HMI tags "Standard-Variablentabelle"
   "Trigger" : Int, internal
   "TP_Online" : Int, internal
   "_BildNr_aktuell" : Int, internal
   "__Pult_Name" : Int, internal
   "__Pult_Name(1)" : WString[10], internal
   "test" : Int, internal
   "LinePLC1_RD_ready" : Bool = PLC LinePLC1_RD_ready AT %I4248.0, 1 s
   "DiagStatusUpdate" : Bool = PLC DiagStatusUpdate AT %M1.1, 1 s
   "EMS_Carrier_Spacing" : Int = PLC EMS.Carrier_Spacing, 1 s
   "EMS_Coarse_Decel_Speed" : Word = PLC EMS.CoarseDecelSpeed AT %DB1.DBW0, 1 s
   "EMS_Coarse_Position_Decel_Offset" : Word = PLC EMS.CoarsePositionDecelOffset AT %DB1.DBW0, 1 s
   "EMS_Coarse_Position_Tolerance" : Word = PLC EMS.CoarsePositionTolerance AT %DB1.DBW0, 1 s
   "EMS_Fine_Decel_Speed" : Word = PLC EMS.FineDecelSpeed AT %DB1.DBW0, 1 s
   "EMS_Fine_Posistion_Tolerance" : Word = PLC EMS.FinePositionTolerance AT %DB1.DBW0, 1 s
   "EMS_Fine_Position_Decel_Offset" : Word = PLC EMS.FinePositionDecelOffset AT %DB1.DBW0, 1 s
   "EMS_Production_Spacing" : Word = PLC EMS.Production_Spacing, 1 s
   "EMS_Production_Zone_Speed" : Word = PLC EMS.ProductionZnSpeed AT %DB1.DBW0, 1 s
   "Temp_Placeholder" : Int = PLC Temp_Int AT %MW56, 1 s
   "CARRIER #01   CURRENT" : Int = PLC "CARRIER #01   CURRENT" AT %MW72, 1 s
   "CARRIER #01   G120D Status WORD.0(1)" : Bool = PLC "CARRIER #01   G120D STATUS WORD.0" AT %M76.0, 1 s
   "CARRIER #01   G120D Status WORD.1(1)" : Bool = PLC "CARRIER #01   G120D STATUS WORD.1" AT %M76.1, 1 s
   "CARRIER #01   G120D Status WORD.10(1)" : Bool = PLC "CARRIER #01   G120D STATUS WORD.10" AT %M77.2, 1 s
   "CARRIER #01   G120D Status WORD.11(1)" : Bool = PLC "CARRIER #01   G120D STATUS WORD.11" AT %M77.3, 1 s
   "CARRIER #01   G120D Status WORD.12(1)" : Bool = PLC "CARRIER #01   G120D STATUS WORD.12" AT %M77.4, 1 s
   "CARRIER #01   G120D Status WORD.13(1)" : Bool = PLC "CARRIER #01   G120D STATUS WORD.13" AT %M77.5, 1 s
   "CARRIER #01   G120D Status WORD.14(1)" : Bool = PLC "CARRIER #01   G120D STATUS WORD.14" AT %M77.6, 1 s
   "CARRIER #01   G120D Status WORD.15(1)" : Bool = PLC "CARRIER #01   G120D STATUS WORD.15" AT %M77.7, 1 s
   "CARRIER #01   G120D Status WORD.2(1)" : Bool = PLC "CARRIER #01   G120D STATUS WORD.2" AT %M76.2, 1 s
   "CARRIER #01   G120D Status WORD.3(1)" : Bool = PLC "CARRIER #01   G120D STATUS WORD.3" AT %M76.3, 1 s
   "CARRIER #01   G120D Status WORD.4(1)" : Bool = PLC "CARRIER #01   G120D STATUS WORD.4" AT %M76.4, 1 s
   "CARRIER #01   G120D Status WORD.5(1)" : Bool = PLC "CARRIER #01   G120D STATUS WORD.5" AT %M76.5, 1 s
   "CARRIER #01   G120D Status WORD.6(1)" : Bool = PLC "CARRIER #01   G120D STATUS WORD.6" AT %M76.6, 1 s
   "CARRIER #01   G120D Status WORD.7(1)" : Bool = PLC "CARRIER #01   G120D STATUS WORD.7" AT %M76.7, 1 s
   "CARRIER #01   G120D Status WORD.8(1)" : Bool = PLC "CARRIER #01   G120D STATUS WORD.8" AT %M77.0, 1 s
   "CARRIER #01   G120D Status WORD.9(1)" : Bool = PLC "CARRIER #01   G120D STATUS WORD.9" AT %M77.1, 1 s
   "CARRIER #01   G120D STATUS WORD.0" : Bool = PLC "CARRIER #01   G120D STATUS WORD.0" AT %M76.0, 1 s
   "CARRIER #01   G120D STATUS WORD.1" : Bool = PLC "CARRIER #01   G120D STATUS WORD.1" AT %M76.1, 1 s
   "CARRIER #01   G120D STATUS WORD.10" : Bool = PLC "CARRIER #01   G120D STATUS WORD.10" AT %M77.2, 1 s
   "CARRIER #01   G120D STATUS WORD.11" : Bool = PLC "CARRIER #01   G120D STATUS WORD.11" AT %M77.3, 1 s
   "CARRIER #01   G120D STATUS WORD.12" : Bool = PLC "CARRIER #01   G120D STATUS WORD.12" AT %M77.4, 1 s
   "CARRIER #01   G120D STATUS WORD.13" : Bool = PLC "CARRIER #01   G120D STATUS WORD.13" AT %M77.5, 1 s
   "CARRIER #01   G120D STATUS WORD.14" : Bool = PLC "CARRIER #01   G120D STATUS WORD.14" AT %M77.6, 1 s
   "CARRIER #01   G120D STATUS WORD.15" : Bool = PLC "CARRIER #01   G120D STATUS WORD.15" AT %M77.7, 1 s
   "CARRIER #01   G120D STATUS WORD.2" : Bool = PLC "CARRIER #01   G120D STATUS WORD.2" AT %M76.2, 1 s
   "CARRIER #01   G120D STATUS WORD.3" : Bool = PLC "CARRIER #01   G120D STATUS WORD.3" AT %M76.3, 1 s
   "CARRIER #01   G120D STATUS WORD.4" : Bool = PLC "CARRIER #01   G120D STATUS WORD.4" AT %M76.4, 1 s
   "CARRIER #01   G120D STATUS WORD.5" : Bool = PLC "CARRIER #01   G120D STATUS WORD.5" AT %M76.5, 1 s
   "CARRIER #01   G120D STATUS WORD.6" : Bool = PLC "CARRIER #01   G120D STATUS WORD.6" AT %M76.6, 1 s
   "CARRIER #01   G120D STATUS WORD.7" : Bool = PLC "CARRIER #01   G120D STATUS WORD.7" AT %M76.7, 1 s
   "CARRIER #01   G120D STATUS WORD.8" : Bool = PLC "CARRIER #01   G120D STATUS WORD.8" AT %M77.0, 1 s
   "CARRIER #01   G120D STATUS WORD.9" : Bool = PLC "CARRIER #01   G120D STATUS WORD.9" AT %M77.1, 1 s
   "CARRIER #01   POSITION" : Int = PLC "CARRIER #01   POSITION" AT %MW78, 1 s
   "CARRIER #01 480VPowerOn_MDCB1" : Bool = PLC "CARRIER #01 480VPowerOn_MDCB1" AT %M80.0, 1 s
   "CARRIER #01 CrashDetectSW" : Bool = PLC "CARRIER #01 CrashDetectSW" AT %M80.1, 1 s
   "CARRIER #01 DCsupplyOnPSCB2" : Bool = PLC "CARRIER #01 DCsupplyOnPSCB2" AT %M80.2, 1 s
   "CARRIER #01 FaultLight_LH" : Bool = PLC "CARRIER #01 FaultLight_LH" AT %M80.3, 1 s
   "CARRIER #01 FaultLight_RH" : Bool = PLC "CARRIER #01 FaultLight_RH" AT %M80.4, 1 s
   "Carrier #01 HMI 1 Status0.5(1)" : Bool = PLC "CARRIER #01   1 STATUS [0].5" AT %M80.5, 1 s
   "CARRIER #01 PB1_ProdHoldLH" : Bool = PLC "CARRIER #01 PB1_ProdHoldLH" AT %M80.6, 1 s
   "CARRIER #01 PB2_ResetLH" : Bool = PLC "CARRIER #01 PB2_ResetLH" AT %M80.7, 1 s
   "CARRIER #01 PB3_ProdHoldRH" : Bool = PLC "CARRIER #01 PB3_ProdHoldRH" AT %M81.0, 1 s
   "CARRIER #01 PB4_ResetRH" : Bool = PLC "CARRIER #01 PB4_ResetRH" AT %M81.1, 1 s
   "CARRIER #01 RunLight_LH" : Bool = PLC "CARRIER #01 RunLight_LH" AT %M81.2, 1 s
   "CARRIER #01 RunLight_RH" : Bool = PLC "CARRIER #01 RunLight_RH" AT %M81.3, 1 s
   "CARRIER #01 SitopSelectStatus" : Bool = PLC "CARRIER #01 SitopSelectStatus" AT %M81.4, 1 s
   "CARRIER #01 SpareInput(2_1)" : Bool = PLC "CARRIER #01 SpareInput(2_1)" AT %M81.5, 1 s
   "CARRIER #01 SpareInput(2_2)" : Bool = PLC "CARRIER #01 SpareInput(2_2)" AT %M81.6, 1 s
   "CARRIER #01 SpareInput(2_3)" : Bool = PLC "CARRIER #01 SpareInput(2_3)" AT %M81.7, 1 s
   "CARRIER #01 SpareInput(2_4)" : Bool = PLC "CARRIER #01 SpareInput(2_4)" AT %M82.0, 1 s
   "CARRIER #01 SpareInput(2_5)" : Bool = PLC "CARRIER #01 SpareInput(2_5)" AT %M82.1, 1 s
   "CARRIER #01 SpareInput(2_6)" : Bool = PLC "CARRIER #01 SpareInput(2_6)" AT %M82.2, 1 s
   "CARRIER #01 SpareInput(2_7)" : Bool = PLC "CARRIER #01 SpareInput(2_7)" AT %M82.3, 1 s
   "CARRIER #01 SpareInput(4_1)" : Bool = PLC "CARRIER #01 SpareInput(4_1)" AT %M82.4, 1 s
   "CARRIER #01 SpareInput(4_14)" : Bool = PLC "CARRIER #01 SpareInput(4_14)" AT %M82.5, 1 s
   "CARRIER #01 SpareInput(4_15)" : Bool = PLC "CARRIER #01 SpareInput(4_15)" AT %M82.6, 1 s
   "CARRIER #01 SpareInput(4_16)" : Bool = PLC "CARRIER #01 SpareInput(4_16)" AT %M82.7, 1 s
   "CARRIER #01 SpareInput(4_17)" : Bool = PLC "CARRIER #01 SpareInput(4_17)" AT %M83.0, 1 s
   "CARRIER #01 SpareInput(4_2)" : Bool = PLC "CARRIER #01 SpareInput(4_2)" AT %M83.1, 1 s
   "CARRIER #01 SpareInput(4_5)" : Bool = PLC "CARRIER #01 SpareInput(4_5)" AT %M83.2, 1 s
   "CARRIER #01 SpareInput(4_6)" : Bool = PLC "CARRIER #01 SpareInput(4_6)" AT %M83.3, 1 s
   "CARRIER #01 SpareInput(4_7)" : Bool = PLC "CARRIER #01 SpareInput(4_7)" AT %M83.4, 1 s
   "CARRIER #01 SpareOutput(5_5)" : Bool = PLC "CARRIER #01 SpareOutput(5_5)" AT %M83.5, 1 s
   "CARRIER #01 SpareOutput(5_6)" : Bool = PLC "CARRIER #01 SpareOutput(5_6)" AT %M83.6, 1 s
   "CARRIER #01 SpareOutput(5_7)" : Bool = PLC "CARRIER #01 SpareOutput(5_7)" AT %M83.7, 1 s
   "CARRIER #01 SpareSafetyOutput(3_1)" : Bool = PLC "CARRIER #01 SpareSafetyOutput(3_1)" AT %M84.0, 1 s
   "CARRIER #01 SpareSafetyOutput(3_2)" : Bool = PLC "CARRIER #01 SpareSafetyOutput(3_2)" AT %M84.1, 1 s
   "CARRIER #01 SpareSafetyOutput(3_3)" : Bool = PLC "CARRIER #01 SpareSafetyOutput(3_3)" AT %M84.2, 1 s
   "CARRIER #01 SpareSafetyOutput(3_4)" : Bool = PLC "CARRIER #01 SpareSafetyOutput(3_4)" AT %M84.3, 1 s
   "CARRIER #01 SpareSafetyOutput(3_5)" : Bool = PLC "CARRIER #01 SpareSafetyOutput(3_5)" AT %M84.4, 1 s
   "CARRIER #01 SpareSafetyOutput(3_6)" : Bool = PLC "CARRIER #01 SpareSafetyOutput(3_6)" AT %M84.5, 1 s
   "CARRIER #01 SpareSafetyOutput(3_7)" : Bool = PLC "CARRIER #01 SpareSafetyOutput(3_7)" AT %M84.6, 1 s
   "Carrier #01_ At Command Position" : Bool = PLC DB_SDC_ERRORS_STAT.ER_AKT[49].ER_STAT[1].ERROR AT %M84.7, 1 s
   "Carrier #01_ Carrier in zone" : Int = PLC "Carrier #01_ Carrier in zone" AT %MW86, 1 s
   "Carrier #01_ Next carrier number" : Int = PLC "Carrier #01_ Next carrier number" AT %MW88, 1 s
   "Carrier 1 G120 D Status" : Bool = PLC EMS.Carrier[12].SDC_IN.DriveCommFault AT %I412.1, 1 s
   "Carrier 1 HMI Status" : Bool = PLC "Carrier 1 HMI Status" AT %I412.2, 1 s
   "Carrier 1 PnF Encoder Status" : Bool = PLC "Carrier 1 PnF Encoder Status" AT %I412.0, 1 s
   "Carrier 2  HMI Staus" : Bool = PLC "Carrier 2 HMI Status" AT %I432.2, 1 s
   "Carrier 2 G120 D Status" : Bool = PLC "Carrier 2  Drive Status" AT %I432.1, 1 s
   "Carrier 2 PnF Encoder Status" : Bool = PLC "Carrier 2 PnF Encoder Status" AT %I432.0, 1 s
   "Carrier 3  G120 D Status" : Bool = PLC "Carrier 3  Drive Status" AT %I452.1, 1 s
   "Carrier 3  PnF Encoder Status" : Bool = PLC "Carrier 3 PnF Encoder Status" AT %I452.0, 1 s
   "Carrier 3 HMI Status" : Bool = PLC "Carrier 3 HMI Status" AT %I452.2, 1 s
   "Carrier 4 G120 D Status" : Bool = PLC "Carrier 4  Drive Status" AT %I472.1, 1 s
   "Carrier 4 HMI Status" : Bool = PLC "Carrier 4 HMI Status" AT %I472.2, 1 s
   "Carrier 4 PnF Encoder Status" : Bool = PLC "Carrier 4 PnF Encoder Status" AT %I472.0, 1 s
   "Carrier_Index_HMI" : Int = PLC Carrier_Index_HMI AT %MW70, 1 s
   "Always_OFF_HMI" : Bool, internal
   "Always_ON_HMI" : Bool, internal
   "EMS_Accum_Zone_Speed" : Word = PLC EMS.AccumZnSpeed AT %DB1.DBW0, 1 s
   "PLC_IP_Address" : WString[30], internal
   "DB302_HMI_Faults_Carrier1_Faults_0" : Int = PLC DB302_HMI_Faults.Carrier1_Faults_0 AT %DB1.DBW0, 1 s
   "DB302_HMI_Faults_Carrier1_Faults_1" : Int = PLC DB302_HMI_Faults.Carrier1_Faults_1 AT %DB1.DBW0, 1 s
   "DB302_HMI_Faults_Carrier1_Faults_2" : Int = PLC DB302_HMI_Faults.Carrier1_Faults_2 AT %DB1.DBW0, 1 s
   "DB302_HMI_Faults_Carrier1_Faults_3" : Int = PLC DB302_HMI_Faults.Carrier1_Faults_3 AT %DB1.DBW0, 1 s
   "DB302_HMI_Faults_Carrier10_Faults_0" : Int = PLC DB302_HMI_Faults.Carrier10_Faults_0 AT %DB1.DBW0, 1 s
   "DB302_HMI_Faults_Carrier10_Faults_1" : Int = PLC DB302_HMI_Faults.Carrier10_Faults_1 AT %DB1.DBW0, 1 s
   "DB302_HMI_Faults_Carrier10_Faults_2" : Int = PLC DB302_HMI_Faults.Carrier10_Faults_2 AT %DB1.DBW0, 1 s
   "DB302_HMI_Faults_Carrier10_Faults_3" : Int = PLC DB302_HMI_Faults.Carrier10_Faults_3 AT %DB1.DBW0, 1 s
   "DB302_HMI_Faults_Carrier11_Faults_0" : Int = PLC DB302_HMI_Faults.Carrier11_Faults_0 AT %DB1.DBW0, 1 s
   "DB302_HMI_Faults_Carrier11_Faults_1" : Int = PLC DB302_HMI_Faults.Carrier11_Faults_1 AT %DB1.DBW0, 1 s
   "DB302_HMI_Faults_Carrier11_Faults_2" : Int = PLC DB302_HMI_Faults.Carrier11_Faults_2 AT %DB1.DBW0, 1 s
   "DB302_HMI_Faults_Carrier11_Faults_3" : Int = PLC DB302_HMI_Faults.Carrier11_Faults_3 AT %DB1.DBW0, 1 s
   "DB302_HMI_Faults_Carrier12_Faults_0" : Int = PLC DB302_HMI_Faults.Carrier12_Faults_0 AT %DB1.DBW0, 1 s
   "DB302_HMI_Faults_Carrier12_Faults_1" : Int = PLC DB302_HMI_Faults.Carrier12_Faults_1 AT %DB1.DBW0, 1 s
   "DB302_HMI_Faults_Carrier12_Faults_2" : Int = PLC DB302_HMI_Faults.Carrier12_Faults_2 AT %DB1.DBW0, 1 s
   "DB302_HMI_Faults_Carrier12_Faults_3" : Int = PLC DB302_HMI_Faults.Carrier12_Faults_3 AT %DB1.DBW0, 1 s
   "DB302_HMI_Faults_Carrier13_Faults_0" : Int = PLC DB302_HMI_Faults.Carrier13_Faults_0 AT %DB1.DBW0, 1 s
   "DB302_HMI_Faults_Carrier13_Faults_1" : Int = PLC DB302_HMI_Faults.Carrier13_Faults_1 AT %DB1.DBW0, 1 s
   "DB302_HMI_Faults_Carrier13_Faults_2" : Int = PLC DB302_HMI_Faults.Carrier13_Faults_2 AT %DB1.DBW0, 1 s
   "DB302_HMI_Faults_Carrier13_Faults_3" : Int = PLC DB302_HMI_Faults.Carrier13_Faults_3 AT %DB1.DBW0, 1 s
   "DB302_HMI_Faults_Carrier14_Faults_0" : Int = PLC DB302_HMI_Faults.Carrier14_Faults_0 AT %DB1.DBW0, 1 s
   "DB302_HMI_Faults_Carrier14_Faults_1" : Int = PLC DB302_HMI_Faults.Carrier14_Faults_1 AT %DB1.DBW0, 1 s
   "DB302_HMI_Faults_Carrier14_Faults_2" : Int = PLC DB302_HMI_Faults.Carrier14_Faults_2 AT %DB1.DBW0, 1 s
   "DB302_HMI_Faults_Carrier14_Faults_3" : Int = PLC DB302_HMI_Faults.Carrier14_Faults_3 AT %DB1.DBW0, 1 s
   "DB302_HMI_Faults_Carrier15_Faults_0" : Int = PLC DB302_HMI_Faults.Carrier15_Faults_0 AT %DB1.DBW0, 1 s
   "DB302_HMI_Faults_Carrier15_Faults_1" : Int = PLC DB302_HMI_Faults.Carrier15_Faults_1 AT %DB1.DBW0, 1 s
   "DB302_HMI_Faults_Carrier15_Faults_2" : Int = PLC DB302_HMI_Faults.Carrier15_Faults_2 AT %DB1.DBW0, 1 s
   "DB302_HMI_Faults_Carrier15_Faults_3" : Int = PLC DB302_HMI_Faults.Carrier15_Faults_3 AT %DB1.DBW0, 1 s
   "DB302_HMI_Faults_Carrier16_Faults_0" : Int = PLC DB302_HMI_Faults.Carrier16_Faults_0 AT %DB1.DBW0, 1 s
   "DB302_HMI_Faults_Carrier16_Faults_1" : Int = PLC DB302_HMI_Faults.Carrier16_Faults_1 AT %DB1.DBW0, 1 s
   "DB302_HMI_Faults_Carrier16_Faults_2" : Int = PLC DB302_HMI_Faults.Carrier16_Faults_2 AT %DB1.DBW0, 1 s
   "DB302_HMI_Faults_Carrier16_Faults_3" : Int = PLC DB302_HMI_Faults.Carrier16_Faults_3 AT %DB1.DBW0, 1 s
   "DB302_HMI_Faults_Carrier17_Faults_0" : Int = PLC DB302_HMI_Faults.Carrier17_Faults_0 AT %DB1.DBW0, 1 s
   "DB302_HMI_Faults_Carrier17_Faults_1" : Int = PLC DB302_HMI_Faults.Carrier17_Faults_1 AT %DB1.DBW0, 1 s
   "DB302_HMI_Faults_Carrier17_Faults_2" : Int = PLC DB302_HMI_Faults.Carrier17_Faults_2 AT %DB1.DBW0, 1 s
   "DB302_HMI_Faults_Carrier17_Faults_3" : Int = PLC DB302_HMI_Faults.Carrier17_Faults_3 AT %DB1.DBW0, 1 s
   "DB302_HMI_Faults_Carrier18_Faults_0" : Int = PLC DB302_HMI_Faults.Carrier18_Faults_0 AT %DB1.DBW0, 1 s
   "DB302_HMI_Faults_Carrier18_Faults_1" : Int = PLC DB302_HMI_Faults.Carrier18_Faults_1 AT %DB1.DBW0, 1 s
   "DB302_HMI_Faults_Carrier18_Faults_2" : Int = PLC DB302_HMI_Faults.Carrier18_Faults_2 AT %DB1.DBW0, 1 s
   "DB302_HMI_Faults_Carrier18_Faults_3" : Int = PLC DB302_HMI_Faults.Carrier18_Faults_3 AT %DB1.DBW0, 1 s
   "DB302_HMI_Faults_Carrier19_Faults_0" : Int = PLC DB302_HMI_Faults.Carrier19_Faults_0 AT %DB1.DBW0, 1 s
   "DB302_HMI_Faults_Carrier19_Faults_1" : Int = PLC DB302_HMI_Faults.Carrier19_Faults_1 AT %DB1.DBW0, 1 s
   "DB302_HMI_Faults_Carrier19_Faults_2" : Int = PLC DB302_HMI_Faults.Carrier19_Faults_2 AT %DB1.DBW0, 1 s
   "DB302_HMI_Faults_Carrier19_Faults_3" : Int = PLC DB302_HMI_Faults.Carrier19_Faults_3 AT %DB1.DBW0, 1 s
   "DB302_HMI_Faults_Carrier2_Faults_0" : Int = PLC DB302_HMI_Faults.Carrier2_Faults_0 AT %DB1.DBW0, 1 s
   "DB302_HMI_Faults_Carrier2_Faults_1" : Int = PLC DB302_HMI_Faults.Carrier2_Faults_1 AT %DB1.DBW0, 1 s
   "DB302_HMI_Faults_Carrier2_Faults_2" : Int = PLC DB302_HMI_Faults.Carrier2_Faults_2 AT %DB1.DBW0, 1 s
   "DB302_HMI_Faults_Carrier2_Faults_3" : Int = PLC DB302_HMI_Faults.Carrier2_Faults_3 AT %DB1.DBW0, 1 s
   "DB302_HMI_Faults_Carrier20_Faults_0" : Int = PLC DB302_HMI_Faults.Carrier20_Faults_0 AT %DB1.DBW0, 1 s
   "DB302_HMI_Faults_Carrier20_Faults_1" : Int = PLC DB302_HMI_Faults.Carrier20_Faults_1 AT %DB1.DBW0, 1 s
   "DB302_HMI_Faults_Carrier20_Faults_2" : Int = PLC DB302_HMI_Faults.Carrier20_Faults_2 AT %DB1.DBW0, 1 s
   "DB302_HMI_Faults_Carrier20_Faults_3" : Int = PLC DB302_HMI_Faults.Carrier20_Faults_3 AT %DB1.DBW0, 1 s
   "DB302_HMI_Faults_Carrier21_Faults_0" : Int = PLC DB302_HMI_Faults.Carrier21_Faults_0 AT %DB1.DBW0, 1 s
   "DB302_HMI_Faults_Carrier21_Faults_1" : Int = PLC DB302_HMI_Faults.Carrier21_Faults_1 AT %DB1.DBW0, 1 s
   "DB302_HMI_Faults_Carrier21_Faults_2" : Int = PLC DB302_HMI_Faults.Carrier21_Faults_2 AT %DB1.DBW0, 1 s
   "DB302_HMI_Faults_Carrier21_Faults_3" : Int = PLC DB302_HMI_Faults.Carrier21_Faults_3 AT %DB1.DBW0, 1 s
   "DB302_HMI_Faults_Carrier22_Faults_0" : Int = PLC DB302_HMI_Faults.Carrier22_Faults_0 AT %DB1.DBW0, 1 s
   "DB302_HMI_Faults_Carrier22_Faults_1" : Int = PLC DB302_HMI_Faults.Carrier22_Faults_1 AT %DB1.DBW0, 1 s
   "DB302_HMI_Faults_Carrier22_Faults_2" : Int = PLC DB302_HMI_Faults.Carrier22_Faults_2 AT %DB1.DBW0, 1 s
   "DB302_HMI_Faults_Carrier22_Faults_3" : Int = PLC DB302_HMI_Faults.Carrier22_Faults_3 AT %DB1.DBW0, 1 s
   "DB302_HMI_Faults_Carrier23_Faults_0" : Int = PLC DB302_HMI_Faults.Carrier23_Faults_0 AT %DB1.DBW0, 1 s
   "DB302_HMI_Faults_Carrier23_Faults_1" : Int = PLC DB302_HMI_Faults.Carrier23_Faults_1 AT %DB1.DBW0, 1 s
   "DB302_HMI_Faults_Carrier23_Faults_2" : Int = PLC DB302_HMI_Faults.Carrier23_Faults_2 AT %DB1.DBW0, 1 s
   "DB302_HMI_Faults_Carrier23_Faults_3" : Int = PLC DB302_HMI_Faults.Carrier23_Faults_3 AT %DB1.DBW0, 1 s
   "DB302_HMI_Faults_Carrier24_Faults_0" : Int = PLC DB302_HMI_Faults.Carrier24_Faults_0 AT %DB1.DBW0, 1 s
   "DB302_HMI_Faults_Carrier24_Faults_1" : Int = PLC DB302_HMI_Faults.Carrier24_Faults_1 AT %DB1.DBW0, 1 s
   "DB302_HMI_Faults_Carrier24_Faults_2" : Int = PLC DB302_HMI_Faults.Carrier24_Faults_2 AT %DB1.DBW0, 1 s
   "DB302_HMI_Faults_Carrier24_Faults_3" : Int = PLC DB302_HMI_Faults.Carrier24_Faults_3 AT %DB1.DBW0, 1 s
   "DB302_HMI_Faults_Carrier25_Faults_0" : Int = PLC DB302_HMI_Faults.Carrier25_Faults_0 AT %DB1.DBW0, 1 s
   "DB302_HMI_Faults_Carrier25_Faults_1" : Int = PLC DB302_HMI_Faults.Carrier25_Faults_1 AT %DB1.DBW0, 1 s
   "DB302_HMI_Faults_Carrier25_Faults_2" : Int = PLC DB302_HMI_Faults.Carrier25_Faults_2 AT %DB1.DBW0, 1 s
   "DB302_HMI_Faults_Carrier25_Faults_3" : Int = PLC DB302_HMI_Faults.Carrier25_Faults_3 AT %DB1.DBW0, 1 s
   "DB302_HMI_Faults_Carrier26_Faults_0" : Int = PLC DB302_HMI_Faults.Carrier26_Faults_0 AT %DB1.DBW0, 1 s
   "DB302_HMI_Faults_Carrier26_Faults_1" : Int = PLC DB302_HMI_Faults.Carrier26_Faults_1 AT %DB1.DBW0, 1 s
   "DB302_HMI_Faults_Carrier26_Faults_2" : Int = PLC DB302_HMI_Faults.Carrier26_Faults_2 AT %DB1.DBW0, 1 s
   "DB302_HMI_Faults_Carrier26_Faults_3" : Int = PLC DB302_HMI_Faults.Carrier26_Faults_3 AT %DB1.DBW0, 1 s
   "DB302_HMI_Faults_Carrier27_Faults_0" : Int = PLC DB302_HMI_Faults.Carrier27_Faults_0 AT %DB1.DBW0, 1 s
   "DB302_HMI_Faults_Carrier27_Faults_1" : Int = PLC DB302_HMI_Faults.Carrier27_Faults_1 AT %DB1.DBW0, 1 s
   "DB302_HMI_Faults_Carrier27_Faults_2" : Int = PLC DB302_HMI_Faults.Carrier27_Faults_2 AT %DB1.DBW0, 1 s
   "DB302_HMI_Faults_Carrier27_Faults_3" : Int = PLC DB302_HMI_Faults.Carrier27_Faults_3 AT %DB1.DBW0, 1 s
   "DB302_HMI_Faults_Carrier28_Faults_0" : Int = PLC DB302_HMI_Faults.Carrier28_Faults_0 AT %DB1.DBW0, 1 s
   "DB302_HMI_Faults_Carrier28_Faults_1" : Int = PLC DB302_HMI_Faults.Carrier28_Faults_1 AT %DB1.DBW0, 1 s
   "DB302_HMI_Faults_Carrier28_Faults_2" : Int = PLC DB302_HMI_Faults.Carrier28_Faults_2 AT %DB1.DBW0, 1 s
   "DB302_HMI_Faults_Carrier28_Faults_3" : Int = PLC DB302_HMI_Faults.Carrier28_Faults_3 AT %DB1.DBW0, 1 s
   "DB302_HMI_Faults_Carrier29_Faults_0" : Int = PLC DB302_HMI_Faults.Carrier29_Faults_0 AT %DB1.DBW0, 1 s
   "DB302_HMI_Faults_Carrier29_Faults_1" : Int = PLC DB302_HMI_Faults.Carrier29_Faults_1 AT %DB1.DBW0, 1 s
   "DB302_HMI_Faults_Carrier29_Faults_2" : Int = PLC DB302_HMI_Faults.Carrier29_Faults_2 AT %DB1.DBW0, 1 s
   "DB302_HMI_Faults_Carrier29_Faults_3" : Int = PLC DB302_HMI_Faults.Carrier29_Faults_3 AT %DB1.DBW0, 1 s
   "DB302_HMI_Faults_Carrier3_Faults_0" : Int = PLC DB302_HMI_Faults.Carrier3_Faults_0 AT %DB1.DBW0, 1 s
   "DB302_HMI_Faults_Carrier3_Faults_1" : Int = PLC DB302_HMI_Faults.Carrier3_Faults_1 AT %DB1.DBW0, 1 s
   "DB302_HMI_Faults_Carrier3_Faults_2" : Int = PLC DB302_HMI_Faults.Carrier3_Faults_2 AT %DB1.DBW0, 1 s
   "DB302_HMI_Faults_Carrier3_Faults_3" : Int = PLC DB302_HMI_Faults.Carrier3_Faults_3 AT %DB1.DBW0, 1 s
   "DB302_HMI_Faults_Carrier30_Faults_0" : Int = PLC DB302_HMI_Faults.Carrier30_Faults_0 AT %DB1.DBW0, 1 s
   "DB302_HMI_Faults_Carrier30_Faults_1" : Int = PLC DB302_HMI_Faults.Carrier30_Faults_1 AT %DB1.DBW0, 1 s
   "DB302_HMI_Faults_Carrier30_Faults_2" : Int = PLC DB_SDC_ERRORS_STAT.ER_AKT[16].ER_STAT[2].DRIVE_POS AT %DB1.DBW0, 1 s
   "DB302_HMI_Faults_Carrier30_Faults_3" : Int = PLC DB302_HMI_Faults.Carrier30_Faults_3 AT %DB1.DBW0, 1 s
   "DB302_HMI_Faults_Carrier31_Faults_0" : Int = PLC DB302_HMI_Faults.Carrier31_Faults_0 AT %DB1.DBW0, 1 s
   "DB302_HMI_Faults_Carrier31_Faults_1" : Int = PLC DB302_HMI_Faults.Carrier31_Faults_1 AT %DB1.DBW0, 1 s
   "DB302_HMI_Faults_Carrier31_Faults_2" : Int = PLC DB302_HMI_Faults.Carrier31_Faults_2 AT %DB1.DBW0, 1 s
   "DB302_HMI_Faults_Carrier31_Faults_3" : Int = PLC DB302_HMI_Faults.Carrier31_Faults_3 AT %DB1.DBW0, 1 s
   "DB302_HMI_Faults_Carrier32_Faults_0" : Int = PLC DB302_HMI_Faults.Carrier32_Faults_0 AT %DB1.DBW0, 1 s
   "DB302_HMI_Faults_Carrier32_Faults_1" : Int = PLC DB302_HMI_Faults.Carrier32_Faults_1 AT %DB1.DBW0, 1 s
   "DB302_HMI_Faults_Carrier32_Faults_2" : Int = PLC DB302_HMI_Faults.Carrier32_Faults_2 AT %DB1.DBW0, 1 s
   "DB302_HMI_Faults_Carrier32_Faults_3" : Int = PLC DB302_HMI_Faults.Carrier32_Faults_3 AT %DB1.DBW0, 1 s
   "DB302_HMI_Faults_Carrier33_Faults_0" : Int = PLC DB302_HMI_Faults.Carrier33_Faults_0 AT %DB1.DBW0, 1 s
   "DB302_HMI_Faults_Carrier33_Faults_1" : Int = PLC DB302_HMI_Faults.Carrier33_Faults_1 AT %DB1.DBW0, 1 s
   "DB302_HMI_Faults_Carrier33_Faults_2" : Int = PLC DB302_HMI_Faults.Carrier33_Faults_2 AT %DB1.DBW0, 1 s
   "DB302_HMI_Faults_Carrier33_Faults_3" : Int = PLC DB302_HMI_Faults.Carrier33_Faults_3 AT %DB1.DBW0, 1 s
   "DB302_HMI_Faults_Carrier34_Faults_0" : Int = PLC DB302_HMI_Faults.Carrier34_Faults_0 AT %DB1.DBW0, 1 s
   "DB302_HMI_Faults_Carrier34_Faults_1" : Int = PLC DB302_HMI_Faults.Carrier34_Faults_1 AT %DB1.DBW0, 1 s
   "DB302_HMI_Faults_Carrier34_Faults_2" : Int = PLC EMS.Carrier[23] AT %DB1.DBW0, 1 s
   "DB302_HMI_Faults_Carrier34_Faults_3" : Int = PLC DB302_HMI_Faults.Carrier34_Faults_3 AT %DB1.DBW0, 1 s
   "DB302_HMI_Faults_Carrier35_Faults_0" : Int = PLC DB302_HMI_Faults.Carrier35_Faults_0 AT %DB1.DBW0, 1 s
   "DB302_HMI_Faults_Carrier35_Faults_1" : Int = PLC DB302_HMI_Faults.Carrier35_Faults_1 AT %DB1.DBW0, 1 s
   "DB302_HMI_Faults_Carrier35_Faults_2" : Int = PLC DB302_HMI_Faults.Carrier35_Faults_2 AT %DB1.DBW0, 1 s
   "DB302_HMI_Faults_Carrier35_Faults_3" : Int = PLC DB302_HMI_Faults.Carrier35_Faults_3 AT %DB1.DBW0, 1 s
   "DB302_HMI_Faults_Carrier36_Faults_0" : Int = PLC DB302_HMI_Faults.Carrier36_Faults_0 AT %DB1.DBW0, 1 s
   "DB302_HMI_Faults_Carrier36_Faults_1" : Int = PLC DB302_HMI_Faults.Carrier36_Faults_1 AT %DB1.DBW0, 1 s
   "DB302_HMI_Faults_Carrier36_Faults_2" : Int = PLC DB302_HMI_Faults.Carrier36_Faults_2 AT %DB1.DBW0, 1 s
   "DB302_HMI_Faults_Carrier36_Faults_3" : Int = PLC DB302_HMI_Faults.Carrier36_Faults_3 AT %DB1.DBW0, 1 s
   "DB302_HMI_Faults_Carrier37_Faults_0" : Int = PLC DB302_HMI_Faults.Carrier37_Faults_0 AT %DB1.DBW0, 1 s
   "DB302_HMI_Faults_Carrier37_Faults_1" : Int = PLC DB302_HMI_Faults.Carrier37_Faults_1 AT %DB1.DBW0, 1 s
   "DB302_HMI_Faults_Carrier37_Faults_2" : Int = PLC DB302_HMI_Faults.Carrier37_Faults_2 AT %DB1.DBW0, 1 s
   "DB302_HMI_Faults_Carrier37_Faults_3" : Int = PLC DB302_HMI_Faults.Carrier37_Faults_3 AT %DB1.DBW0, 1 s
   "DB302_HMI_Faults_Carrier38_Faults_0" : Int = PLC DB302_HMI_Faults.Carrier38_Faults_0 AT %DB1.DBW0, 1 s
   "DB302_HMI_Faults_Carrier38_Faults_1" : Int = PLC DB302_HMI_Faults.Carrier38_Faults_1 AT %DB1.DBW0, 1 s
   "DB302_HMI_Faults_Carrier38_Faults_2" : Int = PLC DB302_HMI_Faults.Carrier38_Faults_2 AT %DB1.DBW0, 1 s
   "DB302_HMI_Faults_Carrier38_Faults_3" : Int = PLC DB302_HMI_Faults.Carrier38_Faults_3 AT %DB1.DBW0, 1 s
   "DB302_HMI_Faults_Carrier39_Faults_0" : Int = PLC DB302_HMI_Faults.Carrier39_Faults_0 AT %DB1.DBW0, 1 s
   "DB302_HMI_Faults_Carrier39_Faults_1" : Int = PLC DB302_HMI_Faults.Carrier39_Faults_1 AT %DB1.DBW0, 1 s
   "DB302_HMI_Faults_Carrier39_Faults_2" : Int = PLC DB302_HMI_Faults.Carrier39_Faults_2 AT %DB1.DBW0, 1 s
   "DB302_HMI_Faults_Carrier39_Faults_3" : Int = PLC DB302_HMI_Faults.Carrier39_Faults_3 AT %DB1.DBW0, 1 s
   "DB302_HMI_Faults_Carrier4_Faults_0" : Int = PLC DB302_HMI_Faults.Carrier4_Faults_0 AT %DB1.DBW0, 1 s
   "DB302_HMI_Faults_Carrier4_Faults_1" : Int = PLC DB302_HMI_Faults.Carrier4_Faults_1 AT %DB1.DBW0, 1 s
   "DB302_HMI_Faults_Carrier4_Faults_2" : Int = PLC DB302_HMI_Faults.Carrier4_Faults_2 AT %DB1.DBW0, 1 s
   "DB302_HMI_Faults_Carrier4_Faults_3" : Int = PLC DB_SDC_BARCODE_INSERTS.INSERT[10].COURSEHIGH AT %DB1.DBW0, 1 s
   "DB302_HMI_Faults_Carrier40_Faults_0" : Int = PLC DB302_HMI_Faults.Carrier40_Faults_0 AT %DB1.DBW0, 1 s
   "DB302_HMI_Faults_Carrier40_Faults_1" : Int = PLC DB302_HMI_Faults.Carrier40_Faults_1 AT %DB1.DBW0, 1 s
   "DB302_HMI_Faults_Carrier40_Faults_2" : Int = PLC DB302_HMI_Faults.Carrier40_Faults_2 AT %DB1.DBW0, 1 s
   "DB302_HMI_Faults_Carrier40_Faults_3" : Int = PLC DB302_HMI_Faults.Carrier40_Faults_3 AT %DB1.DBW0, 1 s
   "DB302_HMI_Faults_Carrier41_Faults_0" : Int = PLC DB302_HMI_Faults.Carrier41_Faults_0 AT %DB1.DBW0, 1 s
   "DB302_HMI_Faults_Carrier41_Faults_1" : Int = PLC DB302_HMI_Faults.Carrier41_Faults_1 AT %DB1.DBW0, 1 s
   "DB302_HMI_Faults_Carrier41_Faults_2" : Int = PLC DB302_HMI_Faults.Carrier41_Faults_2 AT %DB1.DBW0, 1 s
   "DB302_HMI_Faults_Carrier41_Faults_3" : Int = PLC DB302_HMI_Faults.Carrier41_Faults_3 AT %DB1.DBW0, 1 s
   "DB302_HMI_Faults_Carrier42_Faults_0" : Int = PLC DB302_HMI_Faults.Carrier42_Faults_0 AT %DB1.DBW0, 1 s
   "DB302_HMI_Faults_Carrier42_Faults_1" : Int = PLC DB302_HMI_Faults.Carrier42_Faults_1 AT %DB1.DBW0, 1 s
   "DB302_HMI_Faults_Carrier42_Faults_2" : Int = PLC DB302_HMI_Faults.Carrier42_Faults_2 AT %DB1.DBW0, 1 s
   "DB302_HMI_Faults_Carrier42_Faults_3" : Int = PLC DB302_HMI_Faults.Carrier42_Faults_3 AT %DB1.DBW0, 1 s
   "DB302_HMI_Faults_Carrier43_Faults_0" : Int = PLC DB302_HMI_Faults.Carrier43_Faults_0 AT %DB1.DBW0, 1 s
   "DB302_HMI_Faults_Carrier43_Faults_1" : Int = PLC DB302_HMI_Faults.Carrier43_Faults_1 AT %DB1.DBW0, 1 s
   "DB302_HMI_Faults_Carrier43_Faults_2" : Int = PLC DB302_HMI_Faults.Carrier43_Faults_2 AT %DB1.DBW0, 1 s
   "DB302_HMI_Faults_Carrier43_Faults_3" : Int = PLC DB302_HMI_Faults.Carrier43_Faults_3 AT %DB1.DBW0, 1 s
   "DB302_HMI_Faults_Carrier44_Faults_0" : Int = PLC DB302_HMI_Faults.Carrier44_Faults_0 AT %DB1.DBW0, 1 s
   "DB302_HMI_Faults_Carrier44_Faults_1" : Int = PLC DB302_HMI_Faults.Carrier44_Faults_1 AT %DB1.DBW0, 1 s
   "DB302_HMI_Faults_Carrier44_Faults_2" : Int = PLC DB302_HMI_Faults.Carrier44_Faults_2 AT %DB1.DBW0, 1 s
   "DB302_HMI_Faults_Carrier44_Faults_3" : Int = PLC DB302_HMI_Faults.Carrier44_Faults_3 AT %DB1.DBW0, 1 s
   "DB302_HMI_Faults_Carrier45_Faults_0" : Int = PLC DB302_HMI_Faults.Carrier45_Faults_0 AT %DB1.DBW0, 1 s
   "DB302_HMI_Faults_Carrier45_Faults_1" : Int = PLC DB302_HMI_Faults.Carrier45_Faults_1 AT %DB1.DBW0, 1 s
   "DB302_HMI_Faults_Carrier45_Faults_2" : Int = PLC DB302_HMI_Faults.Carrier45_Faults_2 AT %DB1.DBW0, 1 s
   "DB302_HMI_Faults_Carrier45_Faults_3" : Int = PLC DB302_HMI_Faults.Carrier45_Faults_3 AT %DB1.DBW0, 1 s
   "DB302_HMI_Faults_Carrier46_Faults_0" : Int = PLC DB302_HMI_Faults.Carrier46_Faults_0 AT %DB1.DBW0, 1 s
   "DB302_HMI_Faults_Carrier46_Faults_1" : Int = PLC DB302_HMI_Faults.Carrier46_Faults_1 AT %DB1.DBW0, 1 s
   "DB302_HMI_Faults_Carrier46_Faults_2" : Int = PLC DB302_HMI_Faults.Carrier46_Faults_2 AT %DB1.DBW0, 1 s
   "DB302_HMI_Faults_Carrier46_Faults_3" : Int = PLC DB302_HMI_Faults.Carrier46_Faults_3 AT %DB1.DBW0, 1 s
   "DB302_HMI_Faults_Carrier47_Faults_0" : Int = PLC DB302_HMI_Faults.Carrier47_Faults_0 AT %DB1.DBW0, 1 s
   "DB302_HMI_Faults_Carrier47_Faults_1" : Int = PLC DB302_HMI_Faults.Carrier47_Faults_1 AT %DB1.DBW0, 1 s
   "DB302_HMI_Faults_Carrier47_Faults_2" : Int = PLC DB302_HMI_Faults.Carrier47_Faults_2 AT %DB1.DBW0, 1 s
   "DB302_HMI_Faults_Carrier47_Faults_3" : Int = PLC DB302_HMI_Faults.Carrier47_Faults_3 AT %DB1.DBW0, 1 s
   "DB302_HMI_Faults_Carrier48_Faults_0" : Int = PLC DB302_HMI_Faults.Carrier48_Faults_0 AT %DB1.DBW0, 1 s
   "DB302_HMI_Faults_Carrier48_Faults_1" : Int = PLC DB302_HMI_Faults.Carrier48_Faults_1 AT %DB1.DBW0, 1 s
   "DB302_HMI_Faults_Carrier48_Faults_2" : Int = PLC DB302_HMI_Faults.Carrier48_Faults_2 AT %DB1.DBW0, 1 s
   "DB302_HMI_Faults_Carrier48_Faults_3" : Int = PLC DB302_HMI_Faults.Carrier48_Faults_3 AT %DB1.DBW0, 1 s
   "DB302_HMI_Faults_Carrier49_Faults_0" : Int = PLC DB302_HMI_Faults.Carrier49_Faults_0 AT %DB1.DBW0, 1 s
   "DB302_HMI_Faults_Carrier49_Faults_1" : Int = PLC DB302_HMI_Faults.Carrier49_Faults_1 AT %DB1.DBW0, 1 s
   "DB302_HMI_Faults_Carrier49_Faults_2" : Int = PLC DB302_HMI_Faults.Carrier49_Faults_2 AT %DB1.DBW0, 1 s
   "DB302_HMI_Faults_Carrier49_Faults_3" : Int = PLC DB302_HMI_Faults.Carrier49_Faults_3 AT %DB1.DBW0, 1 s
   "DB302_HMI_Faults_Carrier5_Faults_0" : Int = PLC DB302_HMI_Faults.Carrier5_Faults_0 AT %DB1.DBW0, 1 s
   "DB302_HMI_Faults_Carrier5_Faults_1" : Int = PLC DB302_HMI_Faults.Carrier5_Faults_1 AT %DB1.DBW0, 1 s
   "DB302_HMI_Faults_Carrier5_Faults_2" : Int = PLC DB302_HMI_Faults.Carrier5_Faults_2 AT %DB1.DBW0, 1 s
   "DB302_HMI_Faults_Carrier5_Faults_3" : Int = PLC DB302_HMI_Faults.Carrier5_Faults_3 AT %DB1.DBW0, 1 s
   "DB302_HMI_Faults_Carrier50_Faults_0" : Int = PLC DB302_HMI_Faults.Carrier50_Faults_0 AT %DB1.DBW0, 1 s
   "DB302_HMI_Faults_Carrier50_Faults_1" : Int = PLC DB302_HMI_Faults.Carrier50_Faults_1 AT %DB1.DBW0, 1 s
   "DB302_HMI_Faults_Carrier50_Faults_2" : Int = PLC DB302_HMI_Faults.Carrier50_Faults_2 AT %DB1.DBW0, 1 s
   "DB302_HMI_Faults_Carrier50_Faults_3" : Int = PLC DB302_HMI_Faults.Carrier50_Faults_3 AT %DB1.DBW0, 1 s
   "DB302_HMI_Faults_Carrier51_Faults_0" : Int = PLC DB302_HMI_Faults.Carrier51_Faults_0 AT %DB1.DBW0, 1 s
   "DB302_HMI_Faults_Carrier51_Faults_1" : Int = PLC DB302_HMI_Faults.Carrier51_Faults_1 AT %DB1.DBW0, 1 s
   "DB302_HMI_Faults_Carrier51_Faults_2" : Int = PLC DB302_HMI_Faults.Carrier51_Faults_2 AT %DB1.DBW0, 1 s
   "DB302_HMI_Faults_Carrier51_Faults_3" : Int = PLC DB302_HMI_Faults.Carrier51_Faults_3 AT %DB1.DBW0, 1 s